DATA_BLOCK "mst"   // DB33
{ S7_Optimized_Access := 'TRUE' }
VERSION : 0.1
   VAR
      sz : UInt := 9998;
      t : Array[0..10000] of UDInt;
   END_VAR
BEGIN
   t[0] := 1_000_002_001;
   t[1] := 1_000_003_128;
   t[2] := 2_028_513_001;
   t[3] := 33213000;
   t[4] := 2_033_213_010;
   t[5] := 1_033_313_001;
   t[6] := 1_039_413_000;
   t[7] := 2_039_413_010;
   t[8] := 39413011;
   t[9] := 1_039_413_000;
   t[10] := 2_041_813_010;
   t[11] := 41813011;
   t[12] := 2_712_801_002;
   t[13] := 712_801_014;
   t[14] := 712_802_005;
   t[15] := 1_714_701_030;
   t[16] := 1_714_702_014;
   t[17] := 1_714_703_000;
   t[18] := 2_714_701_022;
   t[19] := 2_714_702_010;
   t[20] := 714_701_020;
   t[21] := 1_714_701_016;
   t[22] := 714_901_000;
   t[23] := 714_902_002;
   t[24] := 715_001_016;
   t[25] := 715_002_010;
   t[26] := 1_715_301_000;
   t[27] := 1_715_302_002;
   t[28] := 2_715_401_016;
   t[29] := 2_715_402_010;
   t[30] := 2_715_401_000;
   t[31] := 2_715_402_002;
   t[32] := 715_401_016;
   t[33] := 715_402_010;
   t[34] := 717_702_024;
   t[35] := 717_703_256;
   t[36] := 1_717_702_008;
   t[37] := 1_717_703_000;
   t[38] := 1_717_704_004;
   t[39] := 2_717_703_016;
   t[40] := 717_701_024;
   t[41] := 717_702_012;
   t[42] := 717_703_112;
   t[43] := 718_901_008;
   t[44] := 718_902_004;
   t[45] := 2_719_103_120;
   t[46] := 719_103_121;
   t[47] := 719_203_059;
   t[48] := 1_719_201_000;
   t[49] := 1_719_202_000;
   t[50] := 1_721_203_063;
   t[51] := 2_721_304_008;
   t[52] := 2_721_313_012;
   t[53] := 721_302_001;
   t[54] := 721_303_175;
   t[55] := 721_304_000;
   t[56] := 1_721_303_141;
   t[57] := 723_113_013;
   t[58] := 2_727_713_014;
   t[59] := 1_729_613_015;
   t[60] := 1_733_613_016;
   t[61] := 2_733_612_001;
   t[62] := 736_503_137;
   t[63] := 736_803_129;
   t[64] := 1_736_803_128;
   t[65] := 1_739_013_010;
   t[66] := 2_739_013_011;
   t[67] := 2_741_501_002;
   t[68] := 741_501_014;
   t[69] := 741_502_005;
   t[70] := 2_743_501_030;
   t[71] := 2_743_502_014;
   t[72] := 2_743_503_000;
   t[73] := 743_501_022;
   t[74] := 743_502_010;
   t[75] := 1_743_501_020;
   t[76] := 2_743_501_016;
   t[77] := 743_701_000;
   t[78] := 743_702_002;
   t[79] := 1_743_801_016;
   t[80] := 1_743_802_010;
   t[81] := 746_402_024;
   t[82] := 746_403_256;
   t[83] := 1_746_502_008;
   t[84] := 1_746_503_000;
   t[85] := 1_746_504_004;
   t[86] := 2_746_503_016;
   t[87] := 746_501_024;
   t[88] := 746_502_012;
   t[89] := 746_503_112;
   t[90] := 1_747_501_008;
   t[91] := 1_747_502_004;
   t[92] := 1_747_803_120;
   t[93] := 2_747_803_121;
   t[94] := 2_747_803_059;
   t[95] := 747_801_000;
   t[96] := 747_802_000;
   t[97] := 750_003_063;
   t[98] := 1_750_004_008;
   t[99] := 1_750_013_012;
   t[100] := 2_750_002_001;
   t[101] := 2_750_003_175;
   t[102] := 2_750_004_000;
   t[103] := 750_003_141;
   t[104] := 752_413_013;
   t[105] := 757_013_014;
   t[106] := 2_759_013_015;
   t[107] := 2_763_013_016;
   t[108] := 763_012_002;
   t[109] := 2_766_103_137;
   t[110] := 2_766_303_129;
   t[111] := 766_303_128;
   t[112] := 1_768_613_010;
   t[113] := 2_768_613_011;
   t[114] := 908_001_002;
   t[115] := 1_908_001_014;
   t[116] := 1_908_002_005;
   t[117] := 2_909_901_030;
   t[118] := 2_909_902_014;
   t[119] := 2_909_903_000;
   t[120] := 909_901_022;
   t[121] := 909_902_010;
   t[122] := 1_909_901_020;
   t[123] := 2_909_901_016;
   t[124] := 1_910_001_000;
   t[125] := 1_910_002_002;
   t[126] := 910_201_016;
   t[127] := 910_202_010;
   t[128] := 1_912_902_024;
   t[129] := 1_912_903_256;
   t[130] := 2_912_902_008;
   t[131] := 2_912_903_000;
   t[132] := 2_912_904_004;
   t[133] := 912_903_016;
   t[134] := 1_912_901_024;
   t[135] := 1_912_902_012;
   t[136] := 1_912_903_112;
   t[137] := 1_914_001_008;
   t[138] := 1_914_002_004;
   t[139] := 1_914_303_120;
   t[140] := 2_914_303_121;
   t[141] := 2_914_403_059;
   t[142] := 914_401_000;
   t[143] := 914_402_000;
   t[144] := 2_916_703_063;
   t[145] := 916_704_008;
   t[146] := 916_713_012;
   t[147] := 1_916_702_001;
   t[148] := 1_916_703_175;
   t[149] := 1_916_704_000;
   t[150] := 2_916_703_141;
   t[151] := 1_919_113_013;
   t[152] := 2_923_713_014;
   t[153] := 1_925_713_015;
   t[154] := 2_929_713_016;
   t[155] := 929_712_003;
   t[156] := 1_932_803_137;
   t[157] := 1_933_103_129;
   t[158] := 2_933_103_128;
   t[159] := 1_935_413_010;
   t[160] := 2_935_413_011;
   t[161] := 70547;
   t[162] := 1_160_001_002;
   t[163] := 2_160_001_014;
   t[164] := 2_160_002_005;
   t[165] := 1_161_801_030;
   t[166] := 1_161_802_014;
   t[167] := 1_161_803_000;
   t[168] := 2_161_901_022;
   t[169] := 2_161_902_010;
   t[170] := 161_901_020;
   t[171] := 1_161_901_016;
   t[172] := 162_101_000;
   t[173] := 162_102_002;
   t[174] := 2_162_101_016;
   t[175] := 2_162_102_010;
   t[176] := 1_164_902_024;
   t[177] := 1_164_903_256;
   t[178] := 2_164_902_008;
   t[179] := 2_164_903_000;
   t[180] := 2_164_904_004;
   t[181] := 164_903_016;
   t[182] := 1_164_901_024;
   t[183] := 1_164_902_012;
   t[184] := 1_164_903_112;
   t[185] := 2_166_001_008;
   t[186] := 2_166_002_004;
   t[187] := 1_166_303_120;
   t[188] := 2_166_303_121;
   t[189] := 2_166_303_059;
   t[190] := 166_301_000;
   t[191] := 166_302_000;
   t[192] := 168_603_063;
   t[193] := 1_168_604_008;
   t[194] := 1_168_613_012;
   t[195] := 2_168_602_001;
   t[196] := 2_168_603_175;
   t[197] := 2_168_604_000;
   t[198] := 168_603_141;
   t[199] := 171_013_013;
   t[200] := 2_175_613_014;
   t[201] := 2_177_613_015;
   t[202] := 2_181_713_016;
   t[203] := 181_712_004;
   t[204] := 2_184_603_137;
   t[205] := 185_103_129;
   t[206] := 1_185_103_128;
   t[207] := 187_413_010;
   t[208] := 1_187_413_011;
   t[209] := 205_801_002;
   t[210] := 1_205_801_014;
   t[211] := 1_205_802_005;
   t[212] := 207_701_030;
   t[213] := 207_702_014;
   t[214] := 207_703_000;
   t[215] := 1_207_701_022;
   t[216] := 1_207_702_010;
   t[217] := 2_207_701_020;
   t[218] := 207_701_016;
   t[219] := 2_207_801_000;
   t[220] := 2_207_802_002;
   t[221] := 208_001_016;
   t[222] := 208_002_010;
   t[223] := 2_210_602_024;
   t[224] := 2_210_603_256;
   t[225] := 210_602_008;
   t[226] := 210_603_000;
   t[227] := 210_604_004;
   t[228] := 1_210_603_016;
   t[229] := 2_210_601_024;
   t[230] := 2_210_602_012;
   t[231] := 2_210_603_112;
   t[232] := 1_211_701_008;
   t[233] := 1_211_702_004;
   t[234] := 2_212_003_120;
   t[235] := 212_003_121;
   t[236] := 212_103_059;
   t[237] := 1_212_101_000;
   t[238] := 1_212_102_000;
   t[239] := 2_214_303_063;
   t[240] := 214_304_008;
   t[241] := 214_313_012;
   t[242] := 1_214_302_001;
   t[243] := 1_214_303_175;
   t[244] := 1_214_304_000;
   t[245] := 2_214_303_141;
   t[246] := 2_216_613_013;
   t[247] := 221_313_014;
   t[248] := 2_222_201_002;
   t[249] := 222_201_014;
   t[250] := 222_202_005;
   t[251] := 223_313_015;
   t[252] := 2_224_101_030;
   t[253] := 2_224_102_014;
   t[254] := 2_224_103_013;
   t[255] := 224_101_022;
   t[256] := 224_102_010;
   t[257] := 1_224_101_020;
   t[258] := 2_224_101_016;
   t[259] := 1_227_102_024;
   t[260] := 1_227_103_269;
   t[261] := 227_313_016;
   t[262] := 1_227_312_005;
   t[263] := 1_230_503_265;
   t[264] := 230_803_257;
   t[265] := 1_230_803_256;
   t[266] := 233_113_010;
   t[267] := 1_233_113_011;
   t[268] := 2_234_802_008;
   t[269] := 2_234_803_000;
   t[270] := 2_234_804_004;
   t[271] := 234_803_016;
   t[272] := 1_234_801_024;
   t[273] := 1_234_802_012;
   t[274] := 1_234_803_112;
   t[275] := 2_235_901_008;
   t[276] := 2_235_902_004;
   t[277] := 236_203_120;
   t[278] := 1_236_203_121;
   t[279] := 1_236_203_059;
   t[280] := 2_236_301_000;
   t[281] := 2_236_302_000;
   t[282] := 238_503_063;
   t[283] := 1_238_504_008;
   t[284] := 1_238_513_012;
   t[285] := 2_238_502_001;
   t[286] := 2_238_503_175;
   t[287] := 2_238_504_000;
   t[288] := 238_503_141;
   t[289] := 240_813_013;
   t[290] := 1_245_413_014;
   t[291] := 247_413_015;
   t[292] := 1_251_413_016;
   t[293] := 2_251_412_006;
   t[294] := 2_254_603_137;
   t[295] := 1_254_903_129;
   t[296] := 2_254_903_128;
   t[297] := 257_213_010;
   t[298] := 1_257_313_011;
   t[299] := 70606;
   t[300] := 1_650_801_002;
   t[301] := 2_650_901_014;
   t[302] := 2_650_902_005;
   t[303] := 652_701_030;
   t[304] := 652_702_014;
   t[305] := 652_703_000;
   t[306] := 1_652_701_022;
   t[307] := 1_652_702_010;
   t[308] := 2_652_701_020;
   t[309] := 652_701_016;
   t[310] := 1_652_901_000;
   t[311] := 1_652_902_002;
   t[312] := 1_653_001_016;
   t[313] := 1_653_002_010;
   t[314] := 655_602_024;
   t[315] := 655_603_256;
   t[316] := 1_655_602_008;
   t[317] := 1_655_603_000;
   t[318] := 1_655_604_004;
   t[319] := 2_655_603_016;
   t[320] := 655_601_024;
   t[321] := 655_602_012;
   t[322] := 655_603_112;
   t[323] := 2_656_701_008;
   t[324] := 2_656_702_004;
   t[325] := 1_657_003_120;
   t[326] := 2_657_003_121;
   t[327] := 2_657_003_059;
   t[328] := 657_101_000;
   t[329] := 657_102_000;
   t[330] := 1_659_203_063;
   t[331] := 2_659_204_008;
   t[332] := 2_659_213_012;
   t[333] := 659_202_001;
   t[334] := 659_203_175;
   t[335] := 659_204_000;
   t[336] := 1_659_203_141;
   t[337] := 2_661_513_013;
   t[338] := 666_113_014;
   t[339] := 2_668_113_015;
   t[340] := 2_672_113_016;
   t[341] := 672_112_007;
   t[342] := 675_503_137;
   t[343] := 675_703_129;
   t[344] := 1_675_703_128;
   t[345] := 678_013_010;
   t[346] := 1_678_013_011;
   t[347] := 1_874_401_002;
   t[348] := 2_874_401_014;
   t[349] := 2_874_402_005;
   t[350] := 2_876_201_030;
   t[351] := 2_876_202_014;
   t[352] := 2_876_203_000;
   t[353] := 876_201_022;
   t[354] := 876_202_010;
   t[355] := 1_876_201_020;
   t[356] := 2_876_201_016;
   t[357] := 1_876_301_000;
   t[358] := 1_876_302_002;
   t[359] := 1_876_501_016;
   t[360] := 1_876_502_010;
   t[361] := 879_202_024;
   t[362] := 879_203_256;
   t[363] := 1_879_202_008;
   t[364] := 1_879_203_000;
   t[365] := 1_879_204_004;
   t[366] := 2_879_203_016;
   t[367] := 879_201_024;
   t[368] := 879_202_012;
   t[369] := 879_203_112;
   t[370] := 1_880_201_008;
   t[371] := 1_880_202_004;
   t[372] := 880_503_120;
   t[373] := 1_880_503_121;
   t[374] := 1_880_603_059;
   t[375] := 2_880_601_000;
   t[376] := 2_880_602_000;
   t[377] := 2_882_803_063;
   t[378] := 882_804_008;
   t[379] := 882_813_012;
   t[380] := 1_882_802_001;
   t[381] := 1_882_803_175;
   t[382] := 1_882_804_000;
   t[383] := 2_882_803_141;
   t[384] := 1_885_113_013;
   t[385] := 2_889_713_014;
   t[386] := 891_713_015;
   t[387] := 895_713_016;
   t[388] := 1_895_812_008;
   t[389] := 2_899_003_137;
   t[390] := 1_899_403_129;
   t[391] := 2_899_403_128;
   t[392] := 900_201_002;
   t[393] := 1_900_201_014;
   t[394] := 1_900_202_005;
   t[395] := 2_901_713_010;
   t[396] := 901_713_011;
   t[397] := 902_101_030;
   t[398] := 902_102_014;
   t[399] := 902_103_000;
   t[400] := 1_902_101_022;
   t[401] := 1_902_102_010;
   t[402] := 2_902_101_020;
   t[403] := 902_101_016;
   t[404] := 1_905_102_024;
   t[405] := 1_905_103_256;
   t[406] := 2_905_102_008;
   t[407] := 2_905_103_000;
   t[408] := 2_905_104_004;
   t[409] := 905_103_016;
   t[410] := 1_905_101_024;
   t[411] := 1_905_102_012;
   t[412] := 1_905_103_112;
   t[413] := 906_201_008;
   t[414] := 906_202_004;
   t[415] := 906_403_120;
   t[416] := 1_906_403_121;
   t[417] := 1_906_503_059;
   t[418] := 2_906_501_000;
   t[419] := 2_906_502_000;
   t[420] := 1_908_603_063;
   t[421] := 2_908_604_008;
   t[422] := 2_908_613_012;
   t[423] := 908_602_001;
   t[424] := 908_603_175;
   t[425] := 908_604_000;
   t[426] := 1_908_603_141;
   t[427] := 910_913_013;
   t[428] := 915_613_014;
   t[429] := 2_917_613_015;
   t[430] := 1_921_613_016;
   t[431] := 2_921_612_009;
   t[432] := 924_903_137;
   t[433] := 1_925_203_129;
   t[434] := 2_925_203_128;
   t[435] := 1_927_613_010;
   t[436] := 2_927_613_011;
   t[437] := 1_937_101_002;
   t[438] := 2_937_101_014;
   t[439] := 2_937_102_005;
   t[440] := 2_939_001_030;
   t[441] := 2_939_002_014;
   t[442] := 2_939_003_000;
   t[443] := 939_001_022;
   t[444] := 939_002_010;
   t[445] := 1_939_001_020;
   t[446] := 2_939_001_016;
   t[447] := 1_939_101_000;
   t[448] := 1_939_102_002;
   t[449] := 2_939_201_016;
   t[450] := 2_939_202_010;
   t[451] := 2_942_002_024;
   t[452] := 2_942_003_256;
   t[453] := 942_002_008;
   t[454] := 942_003_000;
   t[455] := 942_004_004;
   t[456] := 1_942_003_016;
   t[457] := 2_942_001_024;
   t[458] := 2_942_002_012;
   t[459] := 2_942_003_112;
   t[460] := 1_943_101_008;
   t[461] := 1_943_102_004;
   t[462] := 1_943_403_120;
   t[463] := 2_943_403_121;
   t[464] := 2_943_403_059;
   t[465] := 943_401_000;
   t[466] := 943_402_000;
   t[467] := 945_803_063;
   t[468] := 1_945_804_008;
   t[469] := 1_945_813_012;
   t[470] := 2_945_802_001;
   t[471] := 2_945_803_175;
   t[472] := 2_945_804_000;
   t[473] := 945_803_141;
   t[474] := 1_948_113_013;
   t[475] := 2_952_713_014;
   t[476] := 2_954_813_015;
   t[477] := 2_958_813_016;
   t[478] := 958_812_010;
   t[479] := 2_962_203_137;
   t[480] := 962_603_129;
   t[481] := 1_962_603_128;
   t[482] := 1_964_913_010;
   t[483] := 2_964_913_011;
   t[484] := 70626;
   t[485] := 25201002;
   t[486] := 1_025_301_014;
   t[487] := 1_025_302_005;
   t[488] := 1_026_901_030;
   t[489] := 1_026_902_014;
   t[490] := 1_026_903_000;
   t[491] := 2_027_001_022;
   t[492] := 2_027_002_010;
   t[493] := 27001020;
   t[494] := 1_027_001_016;
   t[495] := 2_027_101_000;
   t[496] := 2_027_102_002;
   t[497] := 27201016;
   t[498] := 27202010;
   t[499] := 1_030_002_024;
   t[500] := 1_030_003_256;
   t[501] := 2_030_002_008;
   t[502] := 2_030_003_000;
   t[503] := 2_030_004_004;
   t[504] := 30003016;
   t[505] := 1_030_001_024;
   t[506] := 1_030_002_012;
   t[507] := 1_030_003_112;
   t[508] := 30601008;
   t[509] := 30602004;
   t[510] := 2_030_803_120;
   t[511] := 30903121;
   t[512] := 30903059;
   t[513] := 1_030_901_000;
   t[514] := 1_030_902_000;
   t[515] := 33103063;
   t[516] := 1_033_104_008;
   t[517] := 1_033_113_012;
   t[518] := 2_033_102_001;
   t[519] := 2_033_103_175;
   t[520] := 2_033_104_000;
   t[521] := 33103141;
   t[522] := 1_035_513_013;
   t[523] := 1_040_113_014;
   t[524] := 1_042_113_015;
   t[525] := 2_046_213_016;
   t[526] := 46212011;
   t[527] := 2_049_503_137;
   t[528] := 2_049_803_129;
   t[529] := 49903128;
   t[530] := 2_052_313_010;
   t[531] := 52313011;
   t[532] := 1_333_101_002;
   t[533] := 2_333_101_014;
   t[534] := 2_333_102_005;
   t[535] := 1_334_901_030;
   t[536] := 1_334_902_014;
   t[537] := 1_334_903_000;
   t[538] := 2_334_901_022;
   t[539] := 2_334_902_010;
   t[540] := 334_901_020;
   t[541] := 1_335_001_016;
   t[542] := 335_101_000;
   t[543] := 335_102_002;
   t[544] := 2_335_201_016;
   t[545] := 2_335_202_010;
   t[546] := 2_337_902_024;
   t[547] := 2_337_903_256;
   t[548] := 337_902_008;
   t[549] := 337_903_000;
   t[550] := 337_904_004;
   t[551] := 1_337_903_016;
   t[552] := 2_337_901_024;
   t[553] := 2_337_902_012;
   t[554] := 2_337_903_112;
   t[555] := 2_339_001_008;
   t[556] := 2_339_002_004;
   t[557] := 2_339_303_120;
   t[558] := 339_303_121;
   t[559] := 339_303_059;
   t[560] := 1_339_301_000;
   t[561] := 1_339_302_000;
   t[562] := 1_341_503_063;
   t[563] := 2_341_504_008;
   t[564] := 2_341_513_012;
   t[565] := 341_502_001;
   t[566] := 341_503_175;
   t[567] := 341_504_000;
   t[568] := 1_341_503_141;
   t[569] := 2_343_913_013;
   t[570] := 1_348_513_014;
   t[571] := 350_513_015;
   t[572] := 1_354_613_016;
   t[573] := 2_354_612_012;
   t[574] := 1_358_103_137;
   t[575] := 1_358_503_129;
   t[576] := 2_358_503_128;
   t[577] := 2_360_813_010;
   t[578] := 360_813_011;
   t[579] := 2_453_201_002;
   t[580] := 453_201_014;
   t[581] := 453_202_005;
   t[582] := 1_454_901_030;
   t[583] := 1_454_902_014;
   t[584] := 1_454_903_000;
   t[585] := 2_454_901_022;
   t[586] := 2_454_902_010;
   t[587] := 454_901_020;
   t[588] := 1_455_001_016;
   t[589] := 1_458_002_024;
   t[590] := 1_458_003_256;
   t[591] := 2_458_002_008;
   t[592] := 2_458_003_000;
   t[593] := 2_458_004_004;
   t[594] := 458_003_016;
   t[595] := 1_458_001_024;
   t[596] := 1_458_002_012;
   t[597] := 1_458_003_112;
   t[598] := 1_459_001_008;
   t[599] := 1_459_002_004;
   t[600] := 1_459_303_120;
   t[601] := 2_459_303_121;
   t[602] := 2_459_403_059;
   t[603] := 459_401_000;
   t[604] := 459_402_000;
   t[605] := 461_603_063;
   t[606] := 1_461_604_008;
   t[607] := 1_461_613_012;
   t[608] := 2_461_602_001;
   t[609] := 2_461_603_175;
   t[610] := 2_461_604_000;
   t[611] := 461_603_141;
   t[612] := 2_463_913_013;
   t[613] := 2_468_613_014;
   t[614] := 1_470_613_015;
   t[615] := 2_474_613_016;
   t[616] := 474_612_013;
   t[617] := 2_478_103_137;
   t[618] := 2_478_503_129;
   t[619] := 478_503_128;
   t[620] := 480_913_010;
   t[621] := 1_480_913_011;
   t[622] := 482_413_017;
   t[623] := 2_484_203_136;
   t[624] := 484_203_137;
   t[625] := 1_484_503_141;
   t[626] := 1_486_613_018;
   t[627] := 1_491_204_001;
   t[628] := 2_491_203_173;
   t[629] := 2_491_204_003;
   t[630] := 2_491_210_001;
   t[631] := 2_491_211_013;
   t[632] := 2_491_213_000;
   t[633] := 491_603_169;
   t[634] := 1_492_303_173;
   t[635] := 1_492_403_169;
   t[636] := 2_492_503_161;
   t[637] := 492_503_160;
   t[638] := 2_493_203_164;
   t[639] := 493_203_165;
   t[640] := 1_493_303_161;
   t[641] := 2_493_303_160;
   t[642] := 1_495_904_002;
   t[643] := 2_495_903_128;
   t[644] := 2_495_904_000;
   t[645] := 2_495_913_010;
   t[646] := 495_913_015;
   t[647] := 500_013_016;
   t[648] := 1_500_012_014;
   t[649] := 2_501_303_136;
   t[650] := 501_303_137;
   t[651] := 501_903_129;
   t[652] := 1_501_903_128;
   t[653] := 2_505_413_010;
   t[654] := 505_413_011;
   t[655] := 1_843_901_002;
   t[656] := 2_843_901_014;
   t[657] := 2_843_902_005;
   t[658] := 2_845_701_030;
   t[659] := 2_845_702_014;
   t[660] := 2_845_703_000;
   t[661] := 845_701_022;
   t[662] := 845_702_010;
   t[663] := 1_845_701_020;
   t[664] := 2_845_701_016;
   t[665] := 2_845_901_000;
   t[666] := 2_845_902_002;
   t[667] := 2_846_001_016;
   t[668] := 2_846_002_010;
   t[669] := 848_702_024;
   t[670] := 848_703_256;
   t[671] := 1_848_702_008;
   t[672] := 1_848_703_000;
   t[673] := 1_848_704_004;
   t[674] := 2_848_703_016;
   t[675] := 848_701_024;
   t[676] := 848_702_012;
   t[677] := 848_703_112;
   t[678] := 1_849_801_008;
   t[679] := 1_849_802_004;
   t[680] := 1_850_003_120;
   t[681] := 2_850_003_121;
   t[682] := 2_850_103_059;
   t[683] := 850_101_000;
   t[684] := 850_102_000;
   t[685] := 2_852_203_063;
   t[686] := 852_204_008;
   t[687] := 852_213_012;
   t[688] := 1_852_202_001;
   t[689] := 1_852_203_175;
   t[690] := 1_852_204_000;
   t[691] := 2_852_303_141;
   t[692] := 2_854_613_013;
   t[693] := 859_313_014;
   t[694] := 861_313_015;
   t[695] := 1_865_313_016;
   t[696] := 2_865_312_015;
   t[697] := 868_203_137;
   t[698] := 2_868_603_129;
   t[699] := 868_603_128;
   t[700] := 870_813_010;
   t[701] := 1_870_813_011;
   t[702] := 1_897_801_002;
   t[703] := 2_897_801_014;
   t[704] := 2_897_802_005;
   t[705] := 1_899_601_030;
   t[706] := 1_899_602_014;
   t[707] := 1_899_603_000;
   t[708] := 2_899_601_022;
   t[709] := 2_899_602_010;
   t[710] := 899_601_020;
   t[711] := 1_899_601_016;
   t[712] := 899_801_000;
   t[713] := 899_802_002;
   t[714] := 1_899_901_016;
   t[715] := 1_899_902_010;
   t[716] := 2_902_602_024;
   t[717] := 2_902_603_256;
   t[718] := 902_602_008;
   t[719] := 902_603_000;
   t[720] := 902_604_004;
   t[721] := 1_902_603_016;
   t[722] := 2_902_701_024;
   t[723] := 2_902_702_012;
   t[724] := 2_902_703_112;
   t[725] := 903_701_008;
   t[726] := 903_702_004;
   t[727] := 904_003_120;
   t[728] := 1_904_003_121;
   t[729] := 1_904_003_059;
   t[730] := 2_904_001_000;
   t[731] := 2_904_002_000;
   t[732] := 906_303_063;
   t[733] := 1_906_404_008;
   t[734] := 1_906_413_012;
   t[735] := 2_906_402_001;
   t[736] := 2_906_403_175;
   t[737] := 2_906_404_000;
   t[738] := 906_403_141;
   t[739] := 1_908_713_013;
   t[740] := 913_313_014;
   t[741] := 2_915_313_015;
   t[742] := 2_919_313_016;
   t[743] := 919_312_016;
   t[744] := 2_922_203_137;
   t[745] := 1_922_603_129;
   t[746] := 2_922_603_128;
   t[747] := 2_924_913_010;
   t[748] := 925_013_011;
   t[749] := 70645;
   t[750] := 80701002;
   t[751] := 1_080_701_014;
   t[752] := 1_080_702_005;
   t[753] := 1_082_501_030;
   t[754] := 1_082_502_014;
   t[755] := 1_082_503_000;
   t[756] := 2_082_501_022;
   t[757] := 2_082_502_010;
   t[758] := 82501020;
   t[759] := 1_082_501_016;
   t[760] := 1_085_502_024;
   t[761] := 1_085_503_256;
   t[762] := 2_085_502_008;
   t[763] := 2_085_503_000;
   t[764] := 2_085_504_004;
   t[765] := 85503016;
   t[766] := 1_085_501_024;
   t[767] := 1_085_502_012;
   t[768] := 1_085_503_112;
   t[769] := 86601008;
   t[770] := 86602004;
   t[771] := 86903120;
   t[772] := 1_086_903_121;
   t[773] := 1_087_003_059;
   t[774] := 2_087_001_000;
   t[775] := 2_087_002_000;
   t[776] := 89303063;
   t[777] := 1_089_404_008;
   t[778] := 1_089_413_012;
   t[779] := 2_089_402_001;
   t[780] := 2_089_403_175;
   t[781] := 2_089_404_000;
   t[782] := 89403141;
   t[783] := 1_091_713_013;
   t[784] := 2_096_313_014;
   t[785] := 98313015;
   t[786] := 102_313_016;
   t[787] := 1_102_312_017;
   t[788] := 105_203_137;
   t[789] := 2_105_503_129;
   t[790] := 105_503_128;
   t[791] := 2_107_913_010;
   t[792] := 107_913_011;
   t[793] := 1_310_501_002;
   t[794] := 2_310_501_014;
   t[795] := 2_310_502_005;
   t[796] := 2_312_401_030;
   t[797] := 2_312_402_014;
   t[798] := 2_312_403_000;
   t[799] := 312_401_022;
   t[800] := 312_402_010;
   t[801] := 1_312_401_020;
   t[802] := 2_312_401_016;
   t[803] := 315_402_024;
   t[804] := 315_403_256;
   t[805] := 1_315_402_008;
   t[806] := 1_315_403_000;
   t[807] := 1_315_404_004;
   t[808] := 2_315_403_016;
   t[809] := 315_501_024;
   t[810] := 315_502_012;
   t[811] := 315_503_112;
   t[812] := 315_801_008;
   t[813] := 315_802_004;
   t[814] := 1_316_103_120;
   t[815] := 2_316_203_121;
   t[816] := 2_316_203_059;
   t[817] := 316_201_000;
   t[818] := 316_202_000;
   t[819] := 2_318_503_063;
   t[820] := 318_504_008;
   t[821] := 318_513_012;
   t[822] := 1_318_502_001;
   t[823] := 1_318_503_175;
   t[824] := 1_318_504_000;
   t[825] := 2_318_503_141;
   t[826] := 1_320_813_013;
   t[827] := 2_325_413_014;
   t[828] := 1_327_413_015;
   t[829] := 1_331_413_016;
   t[830] := 2_331_412_018;
   t[831] := 1_334_403_137;
   t[832] := 334_703_129;
   t[833] := 1_334_703_128;
   t[834] := 1_337_113_010;
   t[835] := 2_337_113_011;
   t[836] := 398_501_002;
   t[837] := 1_398_501_014;
   t[838] := 1_398_502_005;
   t[839] := 400_301_030;
   t[840] := 400_302_014;
   t[841] := 400_303_000;
   t[842] := 1_400_301_022;
   t[843] := 1_400_302_010;
   t[844] := 2_400_301_020;
   t[845] := 400_301_016;
   t[846] := 400_501_000;
   t[847] := 400_502_002;
   t[848] := 400_501_016;
   t[849] := 400_502_010;
   t[850] := 403_302_024;
   t[851] := 403_303_256;
   t[852] := 1_403_402_008;
   t[853] := 1_403_403_000;
   t[854] := 1_403_404_004;
   t[855] := 2_403_403_016;
   t[856] := 403_401_024;
   t[857] := 403_402_012;
   t[858] := 403_403_112;
   t[859] := 404_401_008;
   t[860] := 404_402_004;
   t[861] := 2_404_703_120;
   t[862] := 404_703_121;
   t[863] := 404_803_059;
   t[864] := 1_404_801_000;
   t[865] := 1_404_802_000;
   t[866] := 407_103_063;
   t[867] := 1_407_104_008;
   t[868] := 1_407_113_012;
   t[869] := 2_407_102_001;
   t[870] := 2_407_103_175;
   t[871] := 2_407_104_000;
   t[872] := 407_103_141;
   t[873] := 409_513_013;
   t[874] := 414_113_014;
   t[875] := 2_416_013_015;
   t[876] := 420_113_016;
   t[877] := 1_420_112_019;
   t[878] := 423_103_137;
   t[879] := 2_423_403_129;
   t[880] := 423_403_128;
   t[881] := 425_813_010;
   t[882] := 1_425_813_011;
   t[883] := 1_602_401_002;
   t[884] := 2_602_401_014;
   t[885] := 2_602_402_005;
   t[886] := 1_604_001_030;
   t[887] := 1_604_002_014;
   t[888] := 1_604_003_000;
   t[889] := 2_604_101_022;
   t[890] := 2_604_102_010;
   t[891] := 604_101_020;
   t[892] := 1_604_101_016;
   t[893] := 2_607_002_024;
   t[894] := 2_607_003_256;
   t[895] := 607_002_008;
   t[896] := 607_003_000;
   t[897] := 607_004_004;
   t[898] := 1_607_003_016;
   t[899] := 2_607_001_024;
   t[900] := 2_607_002_012;
   t[901] := 2_607_003_112;
   t[902] := 2_607_901_008;
   t[903] := 2_607_902_004;
   t[904] := 607_901_024;
   t[905] := 607_902_012;
   t[906] := 2_608_201_008;
   t[907] := 2_608_202_004;
   t[908] := 2_608_403_120;
   t[909] := 608_503_121;
   t[910] := 608_503_059;
   t[911] := 1_608_501_000;
   t[912] := 1_608_502_000;
   t[913] := 2_610_603_063;
   t[914] := 610_704_008;
   t[915] := 610_713_012;
   t[916] := 1_610_702_001;
   t[917] := 1_610_703_175;
   t[918] := 1_610_704_000;
   t[919] := 2_610_703_141;
   t[920] := 1_613_013_013;
   t[921] := 617_713_014;
   t[922] := 619_713_015;
   t[923] := 2_623_713_016;
   t[924] := 623_712_020;
   t[925] := 2_626_903_137;
   t[926] := 2_627_403_129;
   t[927] := 627_403_128;
   t[928] := 629_513_010;
   t[929] := 1_629_613_011;
   t[930] := 1_649_101_002;
   t[931] := 2_649_101_014;
   t[932] := 2_649_102_005;
   t[933] := 2_651_001_030;
   t[934] := 2_651_002_014;
   t[935] := 2_651_003_000;
   t[936] := 651_001_022;
   t[937] := 651_002_010;
   t[938] := 1_651_001_020;
   t[939] := 2_651_101_016;
   t[940] := 2_651_201_000;
   t[941] := 2_651_202_002;
   t[942] := 651_401_016;
   t[943] := 651_402_010;
   t[944] := 1_651_601_000;
   t[945] := 1_651_602_002;
   t[946] := 2_651_601_016;
   t[947] := 2_651_602_010;
   t[948] := 1_654_002_024;
   t[949] := 1_654_003_256;
   t[950] := 2_654_102_008;
   t[951] := 2_654_103_000;
   t[952] := 2_654_104_004;
   t[953] := 654_103_016;
   t[954] := 1_654_101_024;
   t[955] := 1_654_102_012;
   t[956] := 1_654_103_112;
   t[957] := 655_201_008;
   t[958] := 655_202_004;
   t[959] := 1_655_403_120;
   t[960] := 2_655_403_121;
   t[961] := 2_655_503_059;
   t[962] := 655_501_000;
   t[963] := 655_502_000;
   t[964] := 1_657_903_063;
   t[965] := 2_657_904_008;
   t[966] := 2_657_913_012;
   t[967] := 657_902_001;
   t[968] := 657_903_175;
   t[969] := 657_904_000;
   t[970] := 1_657_903_141;
   t[971] := 660_313_013;
   t[972] := 2_665_013_014;
   t[973] := 667_013_015;
   t[974] := 1_671_013_016;
   t[975] := 2_671_012_021;
   t[976] := 2_674_303_137;
   t[977] := 1_674_503_129;
   t[978] := 2_674_503_128;
   t[979] := 676_913_010;
   t[980] := 1_676_913_011;
   t[981] := 727_401_002;
   t[982] := 1_727_401_014;
   t[983] := 1_727_402_005;
   t[984] := 1_729_101_030;
   t[985] := 1_729_102_014;
   t[986] := 1_729_103_000;
   t[987] := 2_729_201_022;
   t[988] := 2_729_202_010;
   t[989] := 729_201_020;
   t[990] := 1_729_201_016;
   t[991] := 1_729_301_000;
   t[992] := 1_729_302_002;
   t[993] := 1_729_501_016;
   t[994] := 1_729_502_010;
   t[995] := 732_102_024;
   t[996] := 732_103_256;
   t[997] := 1_732_102_008;
   t[998] := 1_732_103_000;
   t[999] := 1_732_104_004;
   t[1000] := 2_732_103_016;
   t[1001] := 732_101_024;
   t[1002] := 732_102_012;
   t[1003] := 732_103_112;
   t[1004] := 2_733_201_008;
   t[1005] := 2_733_202_004;
   t[1006] := 1_733_503_120;
   t[1007] := 2_733_503_121;
   t[1008] := 2_733_503_059;
   t[1009] := 733_501_000;
   t[1010] := 733_502_000;
   t[1011] := 2_735_703_063;
   t[1012] := 735_704_008;
   t[1013] := 735_713_012;
   t[1014] := 1_735_702_001;
   t[1015] := 1_735_703_175;
   t[1016] := 1_735_704_000;
   t[1017] := 2_735_703_141;
   t[1018] := 1_738_113_013;
   t[1019] := 742_713_014;
   t[1020] := 2_744_713_015;
   t[1021] := 748_813_016;
   t[1022] := 1_748_812_022;
   t[1023] := 2_751_803_137;
   t[1024] := 752_103_129;
   t[1025] := 1_752_103_128;
   t[1026] := 754_713_010;
   t[1027] := 1_754_813_011;
   t[1028] := 70704;
   t[1029] := 22101002;
   t[1030] := 1_022_101_014;
   t[1031] := 1_022_102_005;
   t[1032] := 2_023_901_030;
   t[1033] := 2_023_902_014;
   t[1034] := 2_023_903_000;
   t[1035] := 23901022;
   t[1036] := 23902010;
   t[1037] := 1_023_901_020;
   t[1038] := 2_023_901_016;
   t[1039] := 1_024_201_000;
   t[1040] := 1_024_202_002;
   t[1041] := 2_024_201_016;
   t[1042] := 2_024_202_010;
   t[1043] := 1_026_802_024;
   t[1044] := 1_026_803_256;
   t[1045] := 2_026_802_008;
   t[1046] := 2_026_803_000;
   t[1047] := 2_026_804_004;
   t[1048] := 26803016;
   t[1049] := 1_026_801_024;
   t[1050] := 1_026_802_012;
   t[1051] := 1_026_803_112;
   t[1052] := 1_027_901_008;
   t[1053] := 1_027_902_004;
   t[1054] := 28203120;
   t[1055] := 1_028_203_121;
   t[1056] := 28303059;
   t[1057] := 1_028_301_000;
   t[1058] := 1_028_302_000;
   t[1059] := 1_030_403_063;
   t[1060] := 2_030_404_008;
   t[1061] := 2_030_413_012;
   t[1062] := 30402001;
   t[1063] := 30403175;
   t[1064] := 30404000;
   t[1065] := 1_030_403_141;
   t[1066] := 2_032_713_013;
   t[1067] := 37213014;
   t[1068] := 2_039_113_015;
   t[1069] := 43113016;
   t[1070] := 1_043_112_023;
   t[1071] := 2_046_403_137;
   t[1072] := 46603129;
   t[1073] := 1_046_603_128;
   t[1074] := 2_049_013_010;
   t[1075] := 49013011;
   t[1076] := 2_073_603_001;
   t[1077] := 2_073_605_008;
   t[1078] := 2_073_606_130;
   t[1079] := 2_073_608_002;
   t[1080] := 2_073_610_000;
   t[1081] := 2_073_611_000;
   t[1082] := 2_073_612_000;
   t[1083] := 2_073_613_000;
   t[1084] := 2_073_614_001;
   t[1085] := 86605024;
   t[1086] := 1_086_605_056;
   t[1087] := 1_086_606_131;
   t[1088] := 552;
   t[1089] := 611;
   t[1090] := 631;
   t[1091] := 650;
   t[1092] := 710;
   t[1093] := 729;
   t[1094] := 749;
   t[1095] := 808;
   t[1096] := 828;
   t[1097] := 2_001_802_003;
   t[1098] := 1_004_103_047;
   t[1099] := 4102002;
   t[1100] := 1_004_102_000;
   t[1101] := 1_004_103_013;
   t[1102] := 17112032;
   t[1103] := 2_020_403_009;
   t[1104] := 1_020_803_001;
   t[1105] := 2_020_803_000;
   t[1106] := 1_055_501_002;
   t[1107] := 2_055_501_014;
   t[1108] := 2_055_502_004;
   t[1109] := 2_057_301_030;
   t[1110] := 2_057_302_012;
   t[1111] := 57301022;
   t[1112] := 57302008;
   t[1113] := 1_057_301_020;
   t[1114] := 2_057_301_016;
   t[1115] := 1_057_501_000;
   t[1116] := 1_057_502_000;
   t[1117] := 2_057_601_016;
   t[1118] := 2_057_602_008;
   t[1119] := 1_060_302_009;
   t[1120] := 2_060_301_024;
   t[1121] := 2_060_302_013;
   t[1122] := 2_060_303_096;
   t[1123] := 61401008;
   t[1124] := 61402005;
   t[1125] := 2_061_703_104;
   t[1126] := 61703105;
   t[1127] := 61802007;
   t[1128] := 61803043;
   t[1129] := 1_061_801_000;
   t[1130] := 1_061_802_003;
   t[1131] := 64003047;
   t[1132] := 2_064_002_002;
   t[1133] := 64002000;
   t[1134] := 64003013;
   t[1135] := 77012033;
   t[1136] := 2_080_403_009;
   t[1137] := 1_080_703_001;
   t[1138] := 2_080_703_000;
   t[1139] := 1_136_301_002;
   t[1140] := 2_136_301_014;
   t[1141] := 2_136_302_004;
   t[1142] := 2_138_201_030;
   t[1143] := 2_138_202_012;
   t[1144] := 138_301_022;
   t[1145] := 138_302_008;
   t[1146] := 1_138_301_020;
   t[1147] := 2_138_301_016;
   t[1148] := 1_138_401_000;
   t[1149] := 1_138_402_000;
   t[1150] := 2_138_501_016;
   t[1151] := 2_138_502_008;
   t[1152] := 2_141_302_009;
   t[1153] := 141_301_024;
   t[1154] := 141_302_013;
   t[1155] := 141_303_096;
   t[1156] := 142_301_008;
   t[1157] := 142_302_005;
   t[1158] := 2_142_603_104;
   t[1159] := 142_603_105;
   t[1160] := 142_702_007;
   t[1161] := 142_703_043;
   t[1162] := 1_142_701_000;
   t[1163] := 1_142_702_003;
   t[1164] := 144_803_047;
   t[1165] := 2_144_802_002;
   t[1166] := 144_902_000;
   t[1167] := 144_903_013;
   t[1168] := 1_157_912_034;
   t[1169] := 161_403_009;
   t[1170] := 161_803_001;
   t[1171] := 1_161_803_000;
   t[1172] := 222_601_002;
   t[1173] := 1_222_601_014;
   t[1174] := 1_222_602_004;
   t[1175] := 2_224_501_030;
   t[1176] := 2_224_502_012;
   t[1177] := 224_501_022;
   t[1178] := 224_502_008;
   t[1179] := 1_224_501_020;
   t[1180] := 2_224_501_016;
   t[1181] := 2_224_701_000;
   t[1182] := 2_224_702_000;
   t[1183] := 2_224_801_016;
   t[1184] := 2_224_802_008;
   t[1185] := 227_602_009;
   t[1186] := 1_227_601_024;
   t[1187] := 1_227_602_013;
   t[1188] := 1_227_603_096;
   t[1189] := 228_001_008;
   t[1190] := 228_002_005;
   t[1191] := 1_228_001_024;
   t[1192] := 1_228_002_013;
   t[1193] := 2_228_301_008;
   t[1194] := 2_228_302_005;
   t[1195] := 228_401_024;
   t[1196] := 228_402_013;
   t[1197] := 2_228_601_008;
   t[1198] := 2_228_602_005;
   t[1199] := 2_228_903_104;
   t[1200] := 228_903_105;
   t[1201] := 228_902_007;
   t[1202] := 228_903_043;
   t[1203] := 1_228_901_000;
   t[1204] := 1_228_902_003;
   t[1205] := 1_230_903_035;
   t[1206] := 2_231_003_043;
   t[1207] := 1_231_303_047;
   t[1208] := 231_302_002;
   t[1209] := 1_231_302_000;
   t[1210] := 1_231_303_013;
   t[1211] := 2_244_712_035;
   t[1212] := 2_248_403_009;
   t[1213] := 248_803_001;
   t[1214] := 1_248_903_000;
   t[1215] := 1_256_401_002;
   t[1216] := 2_256_401_014;
   t[1217] := 2_256_402_004;
   t[1218] := 1_258_301_030;
   t[1219] := 1_258_302_012;
   t[1220] := 2_258_301_022;
   t[1221] := 2_258_302_008;
   t[1222] := 258_301_020;
   t[1223] := 1_258_301_016;
   t[1224] := 2_258_501_000;
   t[1225] := 2_258_502_000;
   t[1226] := 1_258_601_016;
   t[1227] := 1_258_602_008;
   t[1228] := 1_261_302_009;
   t[1229] := 2_261_301_024;
   t[1230] := 2_261_302_013;
   t[1231] := 2_261_303_096;
   t[1232] := 262_401_008;
   t[1233] := 262_402_005;
   t[1234] := 1_262_603_104;
   t[1235] := 2_262_603_105;
   t[1236] := 2_262_702_007;
   t[1237] := 2_262_703_043;
   t[1238] := 262_701_000;
   t[1239] := 262_702_003;
   t[1240] := 2_264_803_047;
   t[1241] := 1_264_802_002;
   t[1242] := 2_264_802_000;
   t[1243] := 2_264_803_013;
   t[1244] := 1_277_912_036;
   t[1245] := 1_281_603_009;
   t[1246] := 1_281_903_001;
   t[1247] := 2_281_903_000;
   t[1248] := 1_307_301_002;
   t[1249] := 2_307_301_014;
   t[1250] := 2_307_302_004;
   t[1251] := 2_309_101_030;
   t[1252] := 2_309_102_012;
   t[1253] := 309_101_022;
   t[1254] := 309_102_008;
   t[1255] := 1_309_101_020;
   t[1256] := 2_309_101_016;
   t[1257] := 1_309_301_000;
   t[1258] := 1_309_302_000;
   t[1259] := 1_309_401_016;
   t[1260] := 1_309_402_008;
   t[1261] := 1_312_102_009;
   t[1262] := 2_312_101_024;
   t[1263] := 2_312_102_013;
   t[1264] := 2_312_103_096;
   t[1265] := 1_313_201_008;
   t[1266] := 1_313_202_005;
   t[1267] := 2_313_403_104;
   t[1268] := 313_403_105;
   t[1269] := 313_502_007;
   t[1270] := 313_503_043;
   t[1271] := 1_313_501_000;
   t[1272] := 1_313_502_003;
   t[1273] := 315_703_047;
   t[1274] := 2_315_702_002;
   t[1275] := 315_702_000;
   t[1276] := 315_703_013;
   t[1277] := 1_328_001_002;
   t[1278] := 2_328_001_014;
   t[1279] := 2_328_002_004;
   t[1280] := 2_328_712_037;
   t[1281] := 2_329_801_030;
   t[1282] := 2_329_802_012;
   t[1283] := 329_801_022;
   t[1284] := 329_802_008;
   t[1285] := 1_329_801_020;
   t[1286] := 2_329_801_016;
   t[1287] := 1_330_001_000;
   t[1288] := 1_330_002_000;
   t[1289] := 1_330_101_016;
   t[1290] := 1_330_102_008;
   t[1291] := 2_332_603_009;
   t[1292] := 332_903_001;
   t[1293] := 1_332_903_000;
   t[1294] := 336_902_009;
   t[1295] := 1_337_001_024;
   t[1296] := 1_337_002_013;
   t[1297] := 1_337_003_096;
   t[1298] := 2_338_001_008;
   t[1299] := 2_338_002_005;
   t[1300] := 338_203_104;
   t[1301] := 1_338_203_105;
   t[1302] := 1_338_302_007;
   t[1303] := 1_338_303_043;
   t[1304] := 2_338_301_000;
   t[1305] := 2_338_302_003;
   t[1306] := 340_503_047;
   t[1307] := 2_340_502_002;
   t[1308] := 340_502_000;
   t[1309] := 340_503_013;
   t[1310] := 2_353_512_038;
   t[1311] := 2_357_503_009;
   t[1312] := 1_357_803_001;
   t[1313] := 2_357_803_000;
   t[1314] := 409_501_002;
   t[1315] := 1_409_501_014;
   t[1316] := 1_409_502_004;
   t[1317] := 411_301_030;
   t[1318] := 411_302_012;
   t[1319] := 1_411_401_022;
   t[1320] := 1_411_402_008;
   t[1321] := 2_411_401_020;
   t[1322] := 411_401_016;
   t[1323] := 411_501_000;
   t[1324] := 411_502_000;
   t[1325] := 2_411_601_016;
   t[1326] := 2_411_602_008;
   t[1327] := 414_402_009;
   t[1328] := 1_414_401_024;
   t[1329] := 1_414_402_013;
   t[1330] := 1_414_403_096;
   t[1331] := 1_415_401_008;
   t[1332] := 1_415_402_005;
   t[1333] := 1_415_703_104;
   t[1334] := 2_415_703_105;
   t[1335] := 2_415_802_007;
   t[1336] := 2_415_803_043;
   t[1337] := 415_801_000;
   t[1338] := 415_802_003;
   t[1339] := 1_417_903_047;
   t[1340] := 417_902_002;
   t[1341] := 1_417_902_000;
   t[1342] := 1_417_903_013;
   t[1343] := 1_431_012_039;
   t[1344] := 1_435_203_009;
   t[1345] := 2_435_503_001;
   t[1346] := 435_503_000;
   t[1347] := 1_441_801_002;
   t[1348] := 2_441_801_014;
   t[1349] := 2_441_802_004;
   t[1350] := 2_443_601_030;
   t[1351] := 2_443_602_012;
   t[1352] := 443_601_022;
   t[1353] := 443_602_008;
   t[1354] := 1_443_601_020;
   t[1355] := 2_443_601_016;
   t[1356] := 2_443_801_000;
   t[1357] := 2_443_802_000;
   t[1358] := 2_443_901_016;
   t[1359] := 2_443_902_008;
   t[1360] := 446_602_009;
   t[1361] := 1_446_601_024;
   t[1362] := 1_446_602_013;
   t[1363] := 1_446_603_096;
   t[1364] := 447_701_008;
   t[1365] := 447_702_005;
   t[1366] := 448_003_104;
   t[1367] := 1_448_003_105;
   t[1368] := 1_448_102_007;
   t[1369] := 1_448_103_043;
   t[1370] := 2_448_101_000;
   t[1371] := 2_448_102_003;
   t[1372] := 450_303_047;
   t[1373] := 2_450_302_002;
   t[1374] := 450_302_000;
   t[1375] := 450_303_013;
   t[1376] := 463_412_040;
   t[1377] := 2_467_603_009;
   t[1378] := 467_903_001;
   t[1379] := 1_467_903_000;
   t[1380] := 2_490_701_002;
   t[1381] := 490_701_014;
   t[1382] := 490_702_004;
   t[1383] := 492_601_030;
   t[1384] := 492_602_012;
   t[1385] := 1_492_601_022;
   t[1386] := 1_492_602_008;
   t[1387] := 2_492_601_020;
   t[1388] := 492_601_016;
   t[1389] := 1_492_801_000;
   t[1390] := 1_492_802_000;
   t[1391] := 492_901_016;
   t[1392] := 492_902_008;
   t[1393] := 493_201_000;
   t[1394] := 493_202_000;
   t[1395] := 493_301_016;
   t[1396] := 493_302_008;
   t[1397] := 2_575_412_041;
   t[1398] := 577_503_008;
   t[1399] := 1_577_503_009;
   t[1400] := 1_577_703_013;
   t[1401] := 1_584_503_029;
   t[1402] := 2_584_503_189;
   t[1403] := 584_903_185;
   t[1404] := 1_585_503_189;
   t[1405] := 585_703_181;
   t[1406] := 585_803_177;
   t[1407] := 1_585_803_176;
   t[1408] := 1_586_403_180;
   t[1409] := 2_586_403_181;
   t[1410] := 1_586_603_177;
   t[1411] := 2_586_603_176;
   t[1412] := 589_203_160;
   t[1413] := 1_589_203_000;
   t[1414] := 593_212_042;
   t[1415] := 2_594_503_008;
   t[1416] := 594_503_009;
   t[1417] := 595_203_001;
   t[1418] := 1_595_203_000;
   t[1419] := 598_702_009;
   t[1420] := 1_598_701_024;
   t[1421] := 1_598_702_013;
   t[1422] := 1_598_703_096;
   t[1423] := 1_599_501_008;
   t[1424] := 1_599_502_005;
   t[1425] := 2_599_601_024;
   t[1426] := 2_599_602_013;
   t[1427] := 599_801_008;
   t[1428] := 599_802_005;
   t[1429] := 2_600_103_104;
   t[1430] := 600_103_105;
   t[1431] := 600_102_007;
   t[1432] := 600_103_043;
   t[1433] := 1_600_101_000;
   t[1434] := 1_600_102_003;
   t[1435] := 600_403_035;
   t[1436] := 2_600_503_043;
   t[1437] := 2_602_403_047;
   t[1438] := 1_602_402_002;
   t[1439] := 2_602_402_000;
   t[1440] := 2_602_403_013;
   t[1441] := 1_602_401_002;
   t[1442] := 2_602_401_014;
   t[1443] := 2_602_402_004;
   t[1444] := 604_201_030;
   t[1445] := 604_202_012;
   t[1446] := 1_604_201_022;
   t[1447] := 1_604_202_008;
   t[1448] := 2_604_201_020;
   t[1449] := 604_201_016;
   t[1450] := 604_401_000;
   t[1451] := 604_402_000;
   t[1452] := 2_604_401_016;
   t[1453] := 2_604_402_008;
   t[1454] := 615_412_043;
   t[1455] := 618_503_009;
   t[1456] := 2_618_803_001;
   t[1457] := 618_803_000;
   t[1458] := 1_622_702_009;
   t[1459] := 2_622_701_024;
   t[1460] := 2_622_702_013;
   t[1461] := 2_622_703_096;
   t[1462] := 623_801_008;
   t[1463] := 623_802_005;
   t[1464] := 2_624_103_104;
   t[1465] := 624_103_105;
   t[1466] := 624_102_007;
   t[1467] := 624_103_043;
   t[1468] := 1_624_101_000;
   t[1469] := 1_624_102_003;
   t[1470] := 2_626_303_047;
   t[1471] := 1_626_302_002;
   t[1472] := 2_626_402_000;
   t[1473] := 2_626_403_013;
   t[1474] := 628_101_002;
   t[1475] := 1_628_101_014;
   t[1476] := 1_628_102_004;
   t[1477] := 2_630_001_030;
   t[1478] := 2_630_002_012;
   t[1479] := 630_001_022;
   t[1480] := 630_002_008;
   t[1481] := 1_630_001_020;
   t[1482] := 2_630_001_016;
   t[1483] := 2_630_101_000;
   t[1484] := 2_630_102_000;
   t[1485] := 630_301_016;
   t[1486] := 630_302_008;
   t[1487] := 1_639_512_044;
   t[1488] := 2_642_503_009;
   t[1489] := 2_642_903_001;
   t[1490] := 642_903_000;
   t[1491] := 2_646_902_009;
   t[1492] := 646_901_024;
   t[1493] := 646_902_013;
   t[1494] := 646_903_096;
   t[1495] := 648_001_008;
   t[1496] := 648_002_005;
   t[1497] := 2_648_303_104;
   t[1498] := 648_303_105;
   t[1499] := 648_302_007;
   t[1500] := 648_303_043;
   t[1501] := 1_648_301_000;
   t[1502] := 1_648_302_003;
   t[1503] := 650_503_047;
   t[1504] := 2_650_502_002;
   t[1505] := 650_502_000;
   t[1506] := 650_503_013;
   t[1507] := 2_650_501_002;
   t[1508] := 650_501_014;
   t[1509] := 650_502_004;
   t[1510] := 2_652_401_030;
   t[1511] := 2_652_402_012;
   t[1512] := 652_401_022;
   t[1513] := 652_402_008;
   t[1514] := 1_652_401_020;
   t[1515] := 2_652_401_016;
   t[1516] := 2_652_601_000;
   t[1517] := 2_652_602_000;
   t[1518] := 652_701_016;
   t[1519] := 652_702_008;
   t[1520] := 1_663_512_045;
   t[1521] := 2_666_703_009;
   t[1522] := 2_667_003_001;
   t[1523] := 667_003_000;
   t[1524] := 671_002_009;
   t[1525] := 1_671_001_024;
   t[1526] := 1_671_002_013;
   t[1527] := 1_671_003_096;
   t[1528] := 1_672_101_008;
   t[1529] := 1_672_102_005;
   t[1530] := 1_672_403_104;
   t[1531] := 2_672_403_105;
   t[1532] := 2_672_402_007;
   t[1533] := 2_672_403_043;
   t[1534] := 672_401_000;
   t[1535] := 672_402_003;
   t[1536] := 674_603_047;
   t[1537] := 2_674_602_002;
   t[1538] := 674_602_000;
   t[1539] := 674_603_013;
   t[1540] := 2_687_612_046;
   t[1541] := 690_803_009;
   t[1542] := 1_691_203_001;
   t[1543] := 2_691_203_000;
   t[1544] := 2_732_101_002;
   t[1545] := 732_101_014;
   t[1546] := 732_102_004;
   t[1547] := 734_001_030;
   t[1548] := 734_002_012;
   t[1549] := 1_734_001_022;
   t[1550] := 1_734_002_008;
   t[1551] := 2_734_001_020;
   t[1552] := 734_001_016;
   t[1553] := 2_734_201_000;
   t[1554] := 2_734_202_000;
   t[1555] := 2_734_301_016;
   t[1556] := 2_734_302_008;
   t[1557] := 734_701_000;
   t[1558] := 734_702_000;
   t[1559] := 1_734_701_016;
   t[1560] := 1_734_702_008;
   t[1561] := 737_002_009;
   t[1562] := 1_737_101_024;
   t[1563] := 1_737_102_013;
   t[1564] := 1_737_103_096;
   t[1565] := 1_738_201_008;
   t[1566] := 1_738_202_005;
   t[1567] := 2_738_403_104;
   t[1568] := 738_403_105;
   t[1569] := 738_502_007;
   t[1570] := 738_503_043;
   t[1571] := 1_738_501_000;
   t[1572] := 1_738_502_003;
   t[1573] := 1_740_703_047;
   t[1574] := 740_702_002;
   t[1575] := 1_740_702_000;
   t[1576] := 1_740_703_013;
   t[1577] := 2_753_612_047;
   t[1578] := 756_903_009;
   t[1579] := 2_757_303_001;
   t[1580] := 757_303_000;
   t[1581] := 1_861_101_002;
   t[1582] := 2_861_101_014;
   t[1583] := 2_861_102_004;
   t[1584] := 2_862_901_030;
   t[1585] := 2_862_902_012;
   t[1586] := 862_901_022;
   t[1587] := 862_902_008;
   t[1588] := 1_862_901_020;
   t[1589] := 2_862_901_016;
   t[1590] := 863_101_000;
   t[1591] := 863_102_000;
   t[1592] := 1_863_201_016;
   t[1593] := 1_863_202_008;
   t[1594] := 2_865_902_009;
   t[1595] := 865_901_024;
   t[1596] := 865_902_013;
   t[1597] := 865_903_096;
   t[1598] := 2_867_001_008;
   t[1599] := 2_867_002_005;
   t[1600] := 2_867_303_104;
   t[1601] := 867_303_105;
   t[1602] := 867_402_007;
   t[1603] := 867_403_043;
   t[1604] := 1_867_401_000;
   t[1605] := 1_867_402_003;
   t[1606] := 869_703_047;
   t[1607] := 2_869_702_002;
   t[1608] := 869_702_000;
   t[1609] := 869_703_013;
   t[1610] := 1_882_712_048;
   t[1611] := 1_886_103_009;
   t[1612] := 2_886_403_001;
   t[1613] := 886_403_000;
   t[1614] := 902_601_002;
   t[1615] := 1_902_601_014;
   t[1616] := 1_902_602_004;
   t[1617] := 904_501_030;
   t[1618] := 904_502_012;
   t[1619] := 1_904_501_022;
   t[1620] := 1_904_502_008;
   t[1621] := 2_904_501_020;
   t[1622] := 904_501_016;
   t[1623] := 904_601_000;
   t[1624] := 904_602_000;
   t[1625] := 2_904_701_016;
   t[1626] := 2_904_702_008;
   t[1627] := 907_402_009;
   t[1628] := 1_907_401_024;
   t[1629] := 1_907_402_013;
   t[1630] := 1_907_403_096;
   t[1631] := 1_908_501_008;
   t[1632] := 1_908_502_005;
   t[1633] := 2_908_803_104;
   t[1634] := 908_803_105;
   t[1635] := 908_802_007;
   t[1636] := 908_803_043;
   t[1637] := 1_908_801_000;
   t[1638] := 1_908_802_003;
   t[1639] := 2_911_003_047;
   t[1640] := 1_911_102_002;
   t[1641] := 2_911_102_000;
   t[1642] := 2_911_103_013;
   t[1643] := 2_924_112_049;
   t[1644] := 1_927_603_009;
   t[1645] := 2_927_903_001;
   t[1646] := 927_903_000;
   t[1647] := 929_501_002;
   t[1648] := 1_929_501_014;
   t[1649] := 1_929_502_004;
   t[1650] := 1_931_401_030;
   t[1651] := 1_931_402_012;
   t[1652] := 2_931_401_022;
   t[1653] := 2_931_402_008;
   t[1654] := 931_401_020;
   t[1655] := 1_931_401_016;
   t[1656] := 931_601_000;
   t[1657] := 931_602_000;
   t[1658] := 2_931_701_016;
   t[1659] := 2_931_702_008;
   t[1660] := 934_402_009;
   t[1661] := 1_934_401_024;
   t[1662] := 1_934_402_013;
   t[1663] := 1_934_403_096;
   t[1664] := 935_501_008;
   t[1665] := 935_502_005;
   t[1666] := 2_935_803_104;
   t[1667] := 935_803_105;
   t[1668] := 935_802_007;
   t[1669] := 935_803_043;
   t[1670] := 1_935_801_000;
   t[1671] := 1_935_802_003;
   t[1672] := 1_938_003_047;
   t[1673] := 938_002_002;
   t[1674] := 1_938_002_000;
   t[1675] := 1_938_003_013;
   t[1676] := 951_012_050;
   t[1677] := 954_603_009;
   t[1678] := 1_954_903_001;
   t[1679] := 2_954_903_000;
   t[1680] := 60654;
   t[1681] := 2_111_301_002;
   t[1682] := 111_301_014;
   t[1683] := 111_302_004;
   t[1684] := 2_113_201_030;
   t[1685] := 2_113_202_012;
   t[1686] := 113_201_022;
   t[1687] := 113_202_008;
   t[1688] := 1_113_201_020;
   t[1689] := 2_113_201_016;
   t[1690] := 2_113_301_000;
   t[1691] := 2_113_302_000;
   t[1692] := 113_401_016;
   t[1693] := 113_402_008;
   t[1694] := 2_116_202_009;
   t[1695] := 116_201_024;
   t[1696] := 116_202_013;
   t[1697] := 116_203_096;
   t[1698] := 2_117_301_008;
   t[1699] := 2_117_302_005;
   t[1700] := 117_603_104;
   t[1701] := 1_117_603_105;
   t[1702] := 1_117_602_007;
   t[1703] := 1_117_603_043;
   t[1704] := 2_117_601_000;
   t[1705] := 2_117_602_003;
   t[1706] := 119_803_047;
   t[1707] := 2_119_802_002;
   t[1708] := 119_802_000;
   t[1709] := 119_803_013;
   t[1710] := 1_132_712_051;
   t[1711] := 1_136_503_009;
   t[1712] := 2_136_803_001;
   t[1713] := 136_903_000;
   t[1714] := 1_351_201_002;
   t[1715] := 2_351_201_014;
   t[1716] := 2_351_202_004;
   t[1717] := 353_101_030;
   t[1718] := 353_102_012;
   t[1719] := 1_353_101_022;
   t[1720] := 1_353_102_008;
   t[1721] := 2_353_101_020;
   t[1722] := 353_101_016;
   t[1723] := 2_353_201_000;
   t[1724] := 2_353_202_000;
   t[1725] := 353_301_016;
   t[1726] := 353_302_008;
   t[1727] := 2_356_102_009;
   t[1728] := 356_101_024;
   t[1729] := 356_102_013;
   t[1730] := 356_103_096;
   t[1731] := 2_356_901_008;
   t[1732] := 2_356_902_005;
   t[1733] := 2_357_001_024;
   t[1734] := 2_357_002_013;
   t[1735] := 357_201_008;
   t[1736] := 357_202_005;
   t[1737] := 2_357_503_104;
   t[1738] := 357_503_105;
   t[1739] := 357_502_007;
   t[1740] := 357_503_043;
   t[1741] := 1_357_501_000;
   t[1742] := 1_357_502_003;
   t[1743] := 2_359_703_047;
   t[1744] := 1_359_702_002;
   t[1745] := 2_359_702_000;
   t[1746] := 2_359_703_013;
   t[1747] := 2_372_612_052;
   t[1748] := 2_376_603_009;
   t[1749] := 1_376_803_001;
   t[1750] := 2_376_803_000;
   t[1751] := 2_508_401_002;
   t[1752] := 508_401_014;
   t[1753] := 508_402_004;
   t[1754] := 1_510_401_030;
   t[1755] := 1_510_402_012;
   t[1756] := 2_510_401_022;
   t[1757] := 2_510_402_008;
   t[1758] := 510_401_020;
   t[1759] := 1_510_401_016;
   t[1760] := 1_510_601_000;
   t[1761] := 1_510_602_000;
   t[1762] := 1_510_701_016;
   t[1763] := 1_510_702_008;
   t[1764] := 513_402_009;
   t[1765] := 1_513_401_024;
   t[1766] := 1_513_402_013;
   t[1767] := 1_513_403_096;
   t[1768] := 2_513_901_008;
   t[1769] := 2_513_902_005;
   t[1770] := 1_513_901_024;
   t[1771] := 1_513_902_013;
   t[1772] := 514_201_008;
   t[1773] := 514_202_005;
   t[1774] := 2_514_301_024;
   t[1775] := 2_514_302_013;
   t[1776] := 2_514_401_008;
   t[1777] := 2_514_402_005;
   t[1778] := 1_514_703_104;
   t[1779] := 2_514_703_105;
   t[1780] := 2_514_802_007;
   t[1781] := 2_514_803_043;
   t[1782] := 514_801_000;
   t[1783] := 514_802_003;
   t[1784] := 2_515_103_035;
   t[1785] := 2_515_103_043;
   t[1786] := 2_516_903_047;
   t[1787] := 1_516_902_002;
   t[1788] := 2_516_902_000;
   t[1789] := 2_516_903_013;
   t[1790] := 1_526_801_002;
   t[1791] := 2_526_801_014;
   t[1792] := 2_526_802_004;
   t[1793] := 528_701_030;
   t[1794] := 528_702_012;
   t[1795] := 1_528_701_022;
   t[1796] := 1_528_702_008;
   t[1797] := 2_528_701_020;
   t[1798] := 528_701_016;
   t[1799] := 2_528_901_000;
   t[1800] := 2_528_902_000;
   t[1801] := 529_001_016;
   t[1802] := 529_002_008;
   t[1803] := 529_301_000;
   t[1804] := 529_302_000;
   t[1805] := 1_529_401_016;
   t[1806] := 1_529_402_008;
   t[1807] := 2_529_401_000;